   IOField "I/O field_72" at 566,349 size 60x22; Authorization "Parameter Change"; FormatPattern 9999
      ProcessValue <- "84_Setpoints_PIT402_Main_HighHigh"
   TextField "Text field_38" at 8,349 size 53x22; Text 'IW116'
   IOField "I/O field_29" at 566,511 size 60x22; FormatPattern 9999
   IOField "I/O field_30" at 499,511 size 60x22; FormatPattern 9999
   IOField "I/O field_32" at 361,552 size 60x22; FormatPattern 9999
   IOField "I/O field_33" at 429,552 size 60x22; FormatPattern 9999
   IOField "I/O field_34" at 565,552 size 60x22; FormatPattern 9999
   IOField "I/O field_35" at 498,552 size 60x22; FormatPattern 9999
   TextField "Text field_39" at 1109,687 size 151x62; Text 'To BC Analogue Inputs'
   AlarmView "Alarm view_1" at 0,777 size 1280x23
   TextField "Text field_40" at 23,309 size 1188x123; Text 'Re - Work Required Througout This page'
   Group "Group" at 455,41 size 373x50
   Button "HmiScreenItemData_8" at 469,45 size 355x40; TextOn 'Back'; TextOff 'Text'
   TextField "Screen title" at 455,41 size 373x50; Text 'Screen title'

screen "BC Analogue Outputs" 1280x800, template "Template"
   on GenerateScreen: "TitleUpdater"()
   Button "HmiScreenItemData_1" at 1,1 size 150x43; TextOn 'Back'; TextOff 'Commissioning'
      on Release: ActivateScreen("Commissioning Main Page", 0)
   Button "Button_15" at 34,732 size 100x35; TextOn 'BWTS Digital Inputs'; TextOff 'Back'
      on Click: ActivateScreen("BC Analogue Inputs", 0)
   AlarmView "Alarm view_1" at 0,777 size 1280x23
   TextField "Text field_90" at 750,328 size 64x20; Text 'Reading'
   TextField "Text field_41" at 553,328 size 89x20; Text 'Description'
   TextField "Text field_43" at 437,328 size 37x20; Text 'AO'
   TextField "Text field_52" at 437,295 size 364x26; Text 'Burner Control System PLC (Rack 2)'
   TextField "Text field_4" at 481,444 size 220x22; Text 'Main Fuel Reg Valve Control'
   IOField "I/O field_4" at 749,446 size 70x22; FormatPattern 9999; Unit %
      ProcessValue <- "16_AQ_Data_CV203_CNTRL"
   TextField "Text field_8" at 428,444 size 53x22; Text 'QW100'
   TextField "Text field_9" at 481,368 size 220x22; Text 'Spare'
   TextField "Text field_12" at 480,482 size 220x22; Text 'Main Atom Air Reg Valve Control'
   IOField "I/O field_5" at 749,481 size 70x22; FormatPattern 9999; Unit %
      ProcessValue <- "16_AQ_Data_CV111_CNTRL"
   TextField "Text field_13" at 427,482 size 53x22; Text 'QW102'
   Button "Button_7" at 716,442 size 29x26; TextOff '+'
      on Press: function_b14e0dd5("80_From_HMI_MAN_AQ_INC_100(1)", 0)
      Visibility <- "82_To_HMI_CRNT_MODE_IGG"
   Button "Button_8" at 824,442 size 29x26; TextOff '-'
      on Press: function_b14e0dd5("80_From_HMI_MAN_AQ_DEC_100(1)", 0)
      Visibility <- "82_To_HMI_CRNT_MODE_IGG"
   Button "Button_9" at 716,480 size 29x26; TextOff '+'
      on Press: function_b14e0dd5("80_From_HMI_MAN_AQ_INC_102", 0)
      Visibility <- "82_To_HMI_CRNT_MODE_IGG"
   Button "Button_10" at 824,480 size 29x26; TextOff '-'
      on Press: function_b14e0dd5("80_From_HMI_MAN_AQ_DEC_102", 0)
      Visibility <- "82_To_HMI_CRNT_MODE_IGG"
   Button "Button_11" at 716,364 size 29x26; TextOff '+'
      on Click: SetBit("80_From_HMI_MAN_AQ_INC_96")
      Visibility <- "82_To_HMI_CRNT_MODE_IGG"
   Button "Button_12" at 824,364 size 29x26; TextOff '-'
      on Click: SetBit("80_From_HMI_MAN_AQ_DEC_96")
      Visibility <- "82_To_HMI_CRNT_MODE_IGG"
   Button "Button_13" at 716,405 size 29x26; TextOff '+'
      on Click: SetBit("80_From_HMI_MAN_AQ_INC_98")
      Visibility <- "82_To_HMI_CRNT_MODE_IGG"
   Button "Button_14" at 824,405 size 29x26; TextOff '-'
      on Click: SetBit("80_From_HMI_MAN_AQ_DEC_98")
      Visibility <- "82_To_HMI_CRNT_MODE_IGG"
   IOField "I/O field_6" at 749,368 size 70x22; FormatPattern 9.9; Unit  
      ProcessValue <- "16_AQ_Data_R2_SPR_AQ_96"
   IOField "I/O field_7" at 749,408 size 70x22; FormatPattern 9.9; Unit  
      ProcessValue <- "16_AQ_Data_R2_SPR_AQ_98"
   TextField "Text field_14" at 481,408 size 220x22; Text 'Spare'
   TextField "Text field_15" at 429,368 size 53x22; Text 'QW96'
   TextField "Text field_16" at 428,408 size 53x22; Text 'QW98'
   Group "Group" at 455,41 size 373x50
   Button "HmiScreenItemData_8" at 469,45 size 355x40; TextOn 'Back'; TextOff 'Text'
   TextField "Screen title" at 455,41 size 373x50; Text 'Screen title'

screen "GCU Analogue Outputs" 1280x800, template "Template"
   on GenerateScreen: "TitleUpdater"()
   Button "HmiScreenItemData_1" at 1,1 size 150x43; TextOn 'Back'; TextOff 'Commissioning'
      on Release: ActivateScreen("Commissioning Main Page", 0)
   Button "Button_15" at 34,732 size 100x35; TextOn 'BWTS Digital Inputs'; TextOff 'Back'
      on Click: ActivateScreen("BC Analogue Inputs", 0)
   AlarmView "Alarm view_1" at 0,777 size 1280x23
   TextField "Text field_90" at 750,328 size 64x20; Text 'Reading'
   TextField "Text field_41" at 553,328 size 89x20; Text 'Description'
   TextField "Text field_43" at 437,328 size 37x20; Text 'AO'
   TextField "Text field_52" at 437,295 size 336x26; Text 'GCU Control System PLC (Rack 3)'
   TextField "Text field_4" at 481,444 size 220x22; Text 'Spare'
   IOField "I/O field_4" at 749,446 size 70x22; FormatPattern 9999
      ProcessValue <- "16_AQ_Data_R3_SPR_AQ_804"
   TextField "Text field_8" at 428,444 size 53x22; Text 'QW804'
   TextField "Text field_9" at 481,368 size 220x22; Text 'CV405 GAS VENT POSITION'
   TextField "Text field_12" at 480,482 size 220x22; Text 'Spare'
   IOField "I/O field_5" at 749,481 size 70x22; FormatPattern 9999
      ProcessValue <- "16_AQ_Data_R3_SPR_AQ_806"
   TextField "Text field_13" at 427,482 size 53x22; Text 'QW806'
   Button "Button_7" at 716,442 size 29x26; TextOff '+'
      on Press: function_b14e0dd5("80_From_HMI_MAN_AQ_INC_804", 0)
      Visibility <- "82_To_HMI_CRNT_MODE_GCU"
   Button "Button_8" at 824,442 size 29x26; TextOff '-'
      on Press: function_b14e0dd5("80_From_HMI_MAN_AQ_DEC_804", 0)
      Visibility <- "82_To_HMI_CRNT_MODE_GCU"
   Button "Button_9" at 717,480 size 29x26; TextOff '+'
      on Press: function_b14e0dd5("80_From_HMI_MAN_AQ_INC_806", 0)
      Visibility <- "82_To_HMI_CRNT_MODE_GCU"
   Button "Button_10" at 825,480 size 29x26; TextOff '-'
      on Press: function_b14e0dd5("80_From_HMI_MAN_AQ_DEC_806", 0)
      Visibility <- "82_To_HMI_CRNT_MODE_GCU"
   Button "Button_11" at 716,364 size 29x26; TextOff '+'
      Visibility <- "82_To_HMI_CRNT_MODE_GCU"
      on Press: function_b14e0dd5("80_From_HMI_MAN_AQ_INC_800", 0)
   Button "Button_12" at 824,364 size 29x26; TextOff '-'
      Visibility <- "82_To_HMI_CRNT_MODE_GCU"
      on Press: function_b14e0dd5("80_From_HMI_MAN_AQ_DEC_800", 0)
   Button "Button_13" at 717,405 size 29x26; TextOff '+'
      Visibility <- "82_To_HMI_CRNT_MODE_GCU"
      on Press: function_b14e0dd5("80_From_HMI_MAN_AQ_INC_802", 0)
   Button "Button_14" at 825,405 size 29x26; TextOff '-'
      Visibility <- "82_To_HMI_CRNT_MODE_GCU"
      on Press: function_b14e0dd5("80_From_HMI_MAN_AQ_DEC_802", 0)
   IOField "I/O field_6" at 750,368 size 70x22; FormatPattern 999; Unit   %
      ProcessValue <- "16_AQ_Data_CV405_CNTRL"
   IOField "I/O field_7" at 751,408 size 70x22; FormatPattern 9999; Unit  
      ProcessValue <- "16_AQ_Data_R3_SPR_AQ_802"
   TextField "Text field_14" at 481,408 size 220x22; Text 'Spare'
   TextField "Text field_15" at 429,368 size 53x22; Text 'QW800'
   TextField "Text field_16" at 428,408 size 53x22; Text 'QW802'
   Group "Group" at 455,41 size 373x50
   Button "HmiScreenItemData_8" at 469,45 size 355x40; TextOn 'Back'; TextOff 'Text'
   TextField "Screen title" at 455,41 size 373x50; Text 'Screen title'

screen "BWT Analogue Outputs" 1280x800, template "Template"
   on GenerateScreen: "TitleUpdater"()
   Button "HmiScreenItemData_1" at 1,1 size 150x43; TextOn 'Back'; TextOff 'Commissioning'
      on Release: ActivateScreen("Commissioning Main Page", 0)
   TextField "Text field_90" at 799,171 size 64x20; Text 'Reading'
   TextField "Text field_41" at 602,171 size 89x20; Text 'Description'
   TextField "Text field_43" at 486,171 size 37x20; Text 'AO'
   TextField "Text field_52" at 486,138 size 340x26; Text 'BWT Control System PLC (Rack 3)'
   TextField "Text field_4" at 530,287 size 220x22; Text 'Main Fuel Reg Valve Control'
   IOField "I/O field_4" at 798,289 size 70x22; FormatPattern 9999; Unit %
      ProcessValue <- "16_AQ_Data_CV203_CNTRL"
   TextField "Text field_8" at 477,287 size 53x22; Text 'QW100'
   TextField "Text field_9" at 530,211 size 220x22; Text 'Spare'
   TextField "Text field_12" at 529,325 size 220x22; Text 'Main Atom Air Reg Valve Control'
   IOField "I/O field_5" at 798,324 size 70x22; FormatPattern 9999; Unit %
      ProcessValue <- "16_AQ_Data_CV111_CNTRL"
   TextField "Text field_13" at 476,325 size 53x22; Text 'QW102'
   Button "Button_7" at 765,285 size 29x26; TextOff '+'
      on Press: function_b14e0dd5("80_From_HMI_MAN_AQ_INC_100(1)", 0)
      Visibility <- "82_To_HMI_CRNT_MODE_IGG"
   Button "Button_8" at 873,285 size 29x26; TextOff '-'
      on Press: function_b14e0dd5("80_From_HMI_MAN_AQ_DEC_100(1)", 0)
      Visibility <- "82_To_HMI_CRNT_MODE_IGG"
   Button "Button_9" at 766,323 size 29x26; TextOff '+'
      on Press: function_b14e0dd5("80_From_HMI_MAN_AQ_INC_102", 0)
      Visibility <- "82_To_HMI_CRNT_MODE_IGG"
   Button "Button_10" at 874,323 size 29x26; TextOff '-'
      on Press: function_b14e0dd5("80_From_HMI_MAN_AQ_DEC_102", 0)
      Visibility <- "82_To_HMI_CRNT_MODE_IGG"
   Button "Button_11" at 765,207 size 29x26; TextOff '+'
      on Click: SetBit("80_From_HMI_MAN_AQ_INC_96")
      Visibility <- "82_To_HMI_CRNT_MODE_IGG"
   Button "Button_12" at 873,207 size 29x26; TextOff '-'
      on Click: SetBit("80_From_HMI_MAN_AQ_DEC_96")
      Visibility <- "82_To_HMI_CRNT_MODE_IGG"
   Button "Button_13" at 766,248 size 29x26; TextOff '+'
      on Click: SetBit("80_From_HMI_MAN_AQ_INC_98")
      Visibility <- "82_To_HMI_CRNT_MODE_IGG"
   Button "Button_14" at 874,248 size 29x26; TextOff '-'
      on Click: SetBit("80_From_HMI_MAN_AQ_DEC_98")
      Visibility <- "82_To_HMI_CRNT_MODE_IGG"
   IOField "I/O field_6" at 799,211 size 70x22; FormatPattern 9.9; Unit  
      ProcessValue <- "16_AQ_Data_R2_SPR_AQ_96"
   IOField "I/O field_7" at 800,251 size 70x22; FormatPattern 9.9; Unit  
      ProcessValue <- "16_AQ_Data_R2_SPR_AQ_98"
   TextField "Text field_14" at 530,251 size 220x22; Text 'Spare'
   TextField "Text field_15" at 478,211 size 53x22; Text 'QW96'
   TextField "Text field_16" at 477,251 size 53x22; Text 'QW98'
   Button "Button_15" at 34,732 size 100x35; TextOn 'BWTS Digital Inputs'; TextOff 'Back'
      on Click: ActivateScreen("BC Analogue Inputs", 0)
   AlarmView "Alarm view_1" at 0,777 size 1280x23
   TextField "Text field_1" at 23,309 size 1188x123; Text 'Re - Work Required Througout This page'
   Group "Group" at 455,41 size 373x50
   Button "HmiScreenItemData_8" at 469,45 size 355x40; TextOn 'Back'; TextOff 'Text'
   TextField "Screen title" at 455,41 size 373x50; Text 'Screen title'

screen "BC Target Setpoints" 1280x800, template "Template"
   on GenerateScreen: "TitleUpdater"()
   Button "HmiScreenItemData_1" at 1,1 size 150x43; TextOn 'Back'; TextOff 'Commissioning'
      on Release: ActivateScreen("Commissioning Main Page", 0)
   AlarmView "Alarm view_1" at 0,777 size 1280x23
   TextField "Text field_25" at 394,430 size 407x22; Text 'PIT-113: IGG Main Atom Air Pressure Target'
   TextField "Text field_29" at 814,210 size 68x20; Text 'Setpoint'
   TextField "Text field_33" at 393,468 size 408x22; Text 'PIT-205: IGG Main Fuel Pressure Target'
   IOField "I/O field_58" at 816,468 size 60x22; Authorization "Parameter Change"; FormatPattern 999.99
      ProcessValue <- "84_Setpoints_PIT205_Target(1)"
   TextField "Text field_35" at 394,552 size 406x22; Text 'E-600: O2 Cargo Blanketing Target'
   TextField "Text field_65" at 394,236 size 411x22; Text 'PIT-402: IG Outlet Pressure Pilot Target'
   TextField "Text field_67" at 394,274 size 410x22; Text 'PIT-402: IG Outlet Pressure Main Target'
   TextField "Text field_69" at 395,313 size 407x22; Text 'PIT-402: IG Outlet Pressure Post Target Start'
   TextField "Text field_71" at 395,352 size 406x22; Text 'PIT-402: IG Outlet Pressure Post Target Maximum'
   TextField "Text field_73" at 395,391 size 407x22; Text 'FD-001: Igniter Target'
   TextField "Text field_42" at 394,210 size 89x20; Text 'Description'
   IOField "I/O field_128" at 816,236 size 60x22; Authorization "Parameter Change"; FormatPattern 999.9
      ProcessValue <- "84_Setpoints_PIT402_Pilot_Target(1)"
   IOField "I/O field_133" at 816,274 size 60x22; Authorization "Parameter Change"; FormatPattern 999.9
      ProcessValue <- "84_Setpoints_PIT402_Main_Target(1)"
   IOField "I/O field_138" at 816,313 size 60x22; Authorization "Parameter Change"; FormatPattern 999.9
      ProcessValue <- "84_Setpoints_PIT402_Post_Target_Start"
   IOField "I/O field_53" at 816,430 size 60x22; Authorization "Parameter Change"; FormatPattern 999.9
      ProcessValue <- "84_Setpoints_PIT113_Pilot_Target(1)"
   IOField "I/O field_148" at 816,391 size 60x22; Authorization "Parameter Change"; FormatPattern 999.9
      ProcessValue <- "84_Setpoints_FD001_Min"
   IOField "I/O field_64" at 816,552 size 60x22; Authorization "Parameter Change"; FormatPattern 99.9
      ProcessValue <- "84_Setpoints_E600_CB_Target"
   TextField "Text field_53" at 393,184 size 213x26; Text 'IGG Target Setpoints'
   IOField "I/O field_5" at 815,352 size 60x22; Authorization "Parameter Change"; FormatPattern 999.9
      ProcessValue <- "84_Setpoints_PIT401_Post_Target_Max"
   TextField "Text field_1" at 394,510 size 406x22; Text 'E-600: O2 Ballast Water Treatment Target'
   IOField "I/O field_2" at 816,510 size 60x22; Authorization "Parameter Change"; FormatPattern 9.99
      ProcessValue <- "84_Setpoints_E600_BWT_Target"
   TextField "Text field_2" at 394,595 size 406x22; Text 'PIT-402 Target Ramp Time (s)'
   IOField "I/O field_1" at 816,595 size 60x22; Authorization "Parameter Change"; FormatPattern 99
      ProcessValue <- "19_AUTO_CMNDS_Data_PIT402_Target"
   Group "Group" at 455,41 size 373x50
   Button "HmiScreenItemData_8" at 469,45 size 355x40; TextOn 'Back'; TextOff 'Text'
   TextField "Screen title" at 455,41 size 373x50; Text 'Screen title'

screen "BC Process Times" 1280x800, template "Template"
   on GenerateScreen: "TitleUpdater"()
   Button "HmiScreenItemData_1" at 1,1 size 150x43; TextOn 'Back'; TextOff 'Commissioning'
      on Release: ActivateScreen("Commissioning Main Page", 0)
   Button "Button_1" at 21,736 size 161x32; TextOff 'IGG Step Times'
      on Activate: ActivateScreen("IGG Max Step Times", 0)
   Button "Button_2" at 1091,736 size 161x32; TextOff 'BC Step Times'
      on Activate: ActivateScreen("BC Max Step Times", 0)
   AlarmView "Alarm view_1" at 0,777 size 1280x23
   TextField "Text field_2" at 262,326 size 271x22; Text 'CV114 Open Delay Time'
   TextField "Text field_3" at 551,161 size 65x20; Text 'Time (s)'
   TextField "Text field_4" at 262,354 size 273x22; Text 'CV206 Open Delay Time'
   IOField "I/O field_1" at 546,354 size 60x22; Authorization "Parameter Change"; FormatPattern 999
      ProcessValue <- "86_Times_CV206_OPEN_TIME"
   TextField "Text field_5" at 262,411 size 270x22; Text 'CV215 Open Delay Time'
   TextField "Text field_6" at 262,186 size 272x22; Text 'CV127 Open #1 Delay Time'
   TextField "Text field_7" at 262,214 size 272x22; Text 'CV127 Closed Delay Time'
   TextField "Text field_8" at 262,242 size 271x22; Text 'CV127 Open #2 Delay Time'
   TextField "Text field_9" at 262,270 size 270x22; Text 'CV124 Open Delay Time'
   TextField "Text field_10" at 262,298 size 270x22; Text 'CV124 Close Delay Purge Time'
   TextField "Text field_11" at 262,161 size 89x20; Text 'Description'
   IOField "I/O field_3" at 546,186 size 60x22; Authorization "Parameter Change"; FormatPattern 999
      ProcessValue <- "86_Times_CV127_OPEN_TIME_#1"
   IOField "I/O field_4" at 546,214 size 60x22; Authorization "Parameter Change"; FormatPattern 999
      ProcessValue <- "86_Times_CV127_CLOSED_TIME"
   IOField "I/O field_6" at 546,242 size 60x22; Authorization "Parameter Change"; FormatPattern 999
      ProcessValue <- "86_Times_CV127_OPEN_TIME_#2"
   IOField "I/O field_8" at 546,298 size 60x22; Authorization "Parameter Change"; FormatPattern 999
      ProcessValue <- "86_Times_CV124_CLOSE_TIME_PRG"
   IOField "I/O field_9" at 546,410 size 60x22; Authorization "Parameter Change"; FormatPattern 999
      ProcessValue <- "86_Times_CV215_OPEN_TIME"
   TextField "Text field_12" at 261,135 size 178x26; Text 'BC Process Times'
   IOField "I/O field_10" at 546,270 size 60x22; Authorization "Parameter Change"; FormatPattern 999
      ProcessValue <- "86_Times_CV124_OPEN_TIME"
   TextField "Text field_13" at 262,383 size 270x22; Text 'CV207 Open Delay Time'
   IOField "I/O field_11" at 546,382 size 60x22; Authorization "Parameter Change"; FormatPattern 999
      ProcessValue <- "86_Times_CV207_OPEN_TIME"
   TextField "Text field_17" at 262,439 size 270x22; Text 'CV215 Close Delay Purge Time'
   IOField "I/O field_16" at 546,438 size 60x22; Authorization "Parameter Change"; FormatPattern 999
      ProcessValue <- "86_Times_CV215_CLOSE_TIME_PRG"
   TextField "Text field_18" at 262,467 size 270x22; Text 'CV216 Open Delay Time'
   IOField "I/O field_17" at 546,466 size 60x22; Authorization "Parameter Change"; FormatPattern 999
      ProcessValue <- "86_Times_CV216_OPEN_TIME"
   TextField "Text field_19" at 262,495 size 269x22; Text 'CV216 Close Delay Purge Time'
   IOField "I/O field_18" at 546,494 size 60x22; Authorization "Parameter Change"; FormatPattern 999
      ProcessValue <- "86_Times_CV216_CLOSE_TIME_PRG"
   TextField "Text field_20" at 262,523 size 269x22; Text 'CV216 Open Delay Purge Time'
   IOField "I/O field_19" at 546,522 size 60x22; Authorization "Parameter Change"; FormatPattern 999
      ProcessValue <- "86_Times_CV216_OPEN_TIME_PRG"
   TextField "Text field_21" at 262,552 size 269x22; Text 'CV206 Close Delay Time'
   IOField "I/O field_20" at 546,551 size 60x22; Authorization "Parameter Change"; FormatPattern 999
      ProcessValue <- "86_Times_CV206_CLOSE_TIME"
   TextField "Text field_22" at 636,186 size 269x22; Text 'CV207 Close Delay Time'
   IOField "I/O field_21" at 916,186 size 60x22; Authorization "Parameter Change"; FormatPattern 999
      ProcessValue <- "86_Times_CV207_CLOSE_TIME"
   TextField "Text field_23" at 636,160 size 89x20; Text 'Description'
   TextField "Text field_24" at 923,161 size 65x20; Text 'Time (s)'
   TextField "Text field_26" at 636,214 size 269x22; Text 'CV114 Close Delay Time'
   IOField "I/O field_22" at 916,214 size 60x22; Authorization "Parameter Change"; FormatPattern 999
      ProcessValue <- "86_Times_CV114_CLOSE_TIME"
   TextField "Text field_27" at 636,242 size 269x22; Text 'CV215 Close Delay Time'
   IOField "I/O field_23" at 916,242 size 60x22; Authorization "Parameter Change"; FormatPattern 999
      ProcessValue <- "86_Times_CV215_CLOSE_TIME"
   TextField "Text field_28" at 636,270 size 269x22; Text 'CV216 Close Delay Time'
   IOField "I/O field_24" at 916,270 size 60x22; Authorization "Parameter Change"; FormatPattern 999
      ProcessValue <- "86_Times_CV216_CLOSE_TIME"
   TextField "Text field_30" at 636,298 size 269x22; Text 'CV124 Close Delay Time'
   IOField "I/O field_25" at 916,298 size 60x22; Authorization "Parameter Change"; FormatPattern 999
      ProcessValue <- "86_Times_CV124_CLOSE_TIME"
   TextField "Text field_31" at 636,326 size 269x22; Text 'X001 Maximum Run Time'
   IOField "I/O field_26" at 916,326 size 60x22; Authorization "Parameter Change"; FormatPattern 999
      ProcessValue <- "86_Times_X001_MAX_RUN_TIME"
   TextField "Text field_32" at 636,354 size 269x22; Text 'X001 Run Confirmation Time'
   IOField "I/O field_27" at 916,354 size 60x22; Authorization "Parameter Change"; FormatPattern 999
      ProcessValue <- "86_Times_X001_RUN_CNF_TIME"
   TextField "Text field_34" at 636,383 size 269x22; Text 'Flame Detection Delay'
   IOField "I/O field_28" at 916,382 size 60x22; Authorization "Parameter Change"; FormatPattern 999
      ProcessValue <- "86_Times_FD_DET_DELAY"
   TextField "Text field_36" at 636,411 size 269x22; Text 'Flame Verification Time'
   IOField "I/O field_29" at 916,410 size 60x22; Authorization "Parameter Change"; FormatPattern 999
      ProcessValue <- "86_Times_FD_VRFCTN_TIME"
   TextField "Text field_37" at 636,439 size 269x22; Text 'Flame Detection Time'
   IOField "I/O field_30" at 916,438 size 60x22; Authorization "Parameter Change"; FormatPattern 999
      ProcessValue <- "86_Times_FDU_DET_TIME"
   TextField "Text field_38" at 636,467 size 269x22; Text 'Max Ignition Sequence Run Time'
   IOField "I/O field_31" at 916,466 size 60x22; Authorization "Parameter Change"; FormatPattern 999
      ProcessValue <- "86_Times_MAX_IGNTN_SEQ_TIME"
   TextField "Text field_39" at 636,495 size 269x22; Text 'Max Main Burner Sequence Run Time'
      Visibility <- "AlwaysTRUE"
   IOField "I/O field_32" at 916,494 size 60x22; Authorization "Parameter Change"; FormatPattern 999; Unit h
      ProcessValue <- "86_Times_MAX_MAIN_BURN_SEQ_TIME"
      Visibility <- "AlwaysTRUE"
   TextField "Text field_40" at 636,523 size 269x22; Text 'Max Pilot Burner Purge Sequence Run Time'
   IOField "I/O field_33" at 916,522 size 60x22; Authorization "Parameter Change"; FormatPattern 999
      ProcessValue <- "86_Times_MAX_PILOT_PURGE_SEQ_TIME"
   TextField "Text field_41" at 636,552 size 269x22; Text 'O2 Check Delay Time'
   IOField "I/O field_34" at 916,551 size 60x22; Authorization "Parameter Change"; FormatPattern 999
      ProcessValue <- "86_Times_O2_CHECK_TIME"
   IOField "I/O field_7" at 546,326 size 60x22; Authorization "Parameter Change"; FormatPattern 999
      ProcessValue <- "86_Times_CV114_OPEN_TIME"
   TextField "Text field_43" at 636,582 size 269x22; Text 'Flame Fail Delay'
   IOField "I/O field_35" at 916,581 size 60x22; Authorization "Parameter Change"; FormatPattern 999
      ProcessValue <- "80_From_HMI_FLM_FAIL_DLY"
   Switch "Switch_1" at 987,492 size 32x29; CaptionText 'Switch'; TextOn 'ON'; TextOff 'OFF'; Authorization "User administration"; PictureOff "Design_5_PilotLight_Green_Off"; PictureOn "Design_5_PilotLight_Green_On"
      on Activate: SetBit("80_From_HMI_BurnerProgramedStop")
      ProcessValue <- "80_From_HMI_BurnerProgramedStop"
      Visibility <- "AlwaysTRUE"
   TextField "Text field_44" at 636,613 size 269x22; Text 'FS317 Delayed Fault'
   IOField "I/O field_36" at 916,613 size 60x22; Authorization "Parameter Change"; FormatPattern 999
      ProcessValue <- "86_Times_FS317 delay"
   TextField "Text field_45" at 636,644 size 269x22; Text 'FS320 Delayed Fault'
   IOField "I/O field_37" at 916,644 size 60x22; Authorization "Parameter Change"; FormatPattern 999
      ProcessValue <- "86_Times_FS320 delay"
   TextField "Text field_46" at 262,581 size 269x22; Text 'FS359 Delayed Fault'
   IOField "I/O field_38" at 546,581 size 60x22; Authorization "Parameter Change"; FormatPattern 999
      ProcessValue <- "80_From_HMI_PIT 359 delay"
   TextField "Text field_47" at 262,612 size 269x22; Text 'FS316 Delayed Fault'
   IOField "I/O field_39" at 546,612 size 60x22; Authorization "Parameter Change"; FormatPattern 999
      ProcessValue <- "80_From_HMI_PIT 316 delay"
   Group "Group" at 455,41 size 373x50
   TextField "Text field_1" at 262,643 size 269x22; Text 'PS101 Delayed Fault'
   IOField "I/O field_2" at 546,643 size 60x22; Authorization "Parameter Change"; FormatPattern 999
      ProcessValue <- "86_Times_PS101 Alarm Delay"
   Button "HmiScreenItemData_8" at 469,45 size 355x40; TextOn 'Back'; TextOff 'Text'
   TextField "Screen title" at 455,41 size 373x50; Text 'Screen title'

screen "GCU Max Step Times" 1280x800, template "Template"
   on GenerateScreen: "TitleUpdater"()
   Button "HmiScreenItemData_1" at 1,1 size 150x43; TextOn 'Back'; TextOff 'Commissioning'
      on Release: ActivateScreen("Commissioning Main Page", 0)
   TextField "Text field_29" at 130,95 size 75x25; Text 'Time (ms)'
   TextField "Text field_65" at 40,130 size 75x25; Text 'Step 001'
   TextField "Text field_42" at 40,95 size 75x25; Text 'STEP'
   IOField "I/O field_128" at 130,130 size 75x25; Authorization "Parameter Change"; FormatPattern 999999
      ProcessValue <- "86_Times_STEP_MAX_TIME_STP_001"
   TextField "Text field_53" at 40,66 size 262x26; Text 'GCU Maximum Step Times'
   TextField "Text field_1" at 385,95 size 75x25; Text 'Time (ms)'
   TextField "Text field_2" at 295,130 size 75x25; Text 'Step 170'
   TextField "Text field_3" at 295,95 size 75x25; Text 'STEP'
   IOField "I/O field_1" at 385,130 size 75x25; Authorization "Parameter Change"; FormatPattern 999999
      ProcessValue <- "86_Times_STEP_MAX_TIME_STP_170"
   TextField "Text field_4" at 640,95 size 75x25; Text 'Time (ms)'
   TextField "Text field_5" at 550,130 size 75x25; Text 'Step 350'
   TextField "Text field_6" at 550,95 size 75x25; Text 'STEP'
   IOField "I/O field_2" at 640,130 size 75x25; Authorization "Parameter Change"; FormatPattern 999999
      ProcessValue <- "86_Times_STEP_MAX_TIME_STP_350"
   TextField "Text field_7" at 895,95 size 75x25; Text 'Time (ms)'
   TextField "Text field_8" at 805,130 size 75x25; Text 'Step 530'
   TextField "Text field_9" at 805,95 size 75x25; Text 'STEP'
   IOField "I/O field_3" at 895,130 size 75x25; Authorization "Parameter Change"; FormatPattern 999999
      ProcessValue <- "86_Times_STEP_MAX_TIME_STP_530"
   TextField "Text field_10" at 1150,95 size 75x25; Text 'Time (ms)'
   TextField "Text field_12" at 1060,95 size 75x25; Text 'STEP'
   TextField "Text field_13" at 40,165 size 75x25; Text 'Step 005'
   IOField "I/O field_5" at 130,165 size 75x25; Authorization "Parameter Change"; FormatPattern 999999
      ProcessValue <- "86_Times_STEP_MAX_TIME_STP_005"
   TextField "Text field_14" at 295,165 size 75x25; Text 'Step 180'
   IOField "I/O field_6" at 385,165 size 75x25; Authorization "Parameter Change"; FormatPattern 999999
      ProcessValue <- "86_Times_STEP_MAX_TIME_STP_180"
   TextField "Text field_15" at 550,165 size 75x25; Text 'Step 360'
   IOField "I/O field_7" at 640,165 size 75x25; Authorization "Parameter Change"; FormatPattern 999999
      ProcessValue <- "86_Times_STEP_MAX_TIME_STP_360"
   TextField "Text field_16" at 805,165 size 75x25; Text 'Step 540'
   IOField "I/O field_8" at 895,165 size 75x25; Authorization "Parameter Change"; FormatPattern 999999
      ProcessValue <- "86_Times_STEP_MAX_TIME_STP_540"
   TextField "Text field_18" at 40,200 size 75x25; Text 'Step 010'
   IOField "I/O field_10" at 130,200 size 75x25; Authorization "Parameter Change"; FormatPattern 999999
      ProcessValue <- "86_Times_STEP_MAX_TIME_STP_010"
   TextField "Text field_19" at 295,200 size 75x25; Text 'Step 190'
   IOField "I/O field_11" at 385,200 size 75x25; Authorization "Parameter Change"; FormatPattern 999999
      ProcessValue <- "86_Times_STEP_MAX_TIME_STP_190"
   TextField "Text field_20" at 550,200 size 75x25; Text 'Step 370'
   IOField "I/O field_12" at 640,200 size 75x25; Authorization "Parameter Change"; FormatPattern 999999
      ProcessValue <- "86_Times_STEP_MAX_TIME_STP_370"
   TextField "Text field_21" at 805,200 size 75x25; Text 'Step 550'
   IOField "I/O field_13" at 895,200 size 75x25; Authorization "Parameter Change"; FormatPattern 999999
      ProcessValue <- "86_Times_STEP_MAX_TIME_STP_550"
   TextField "Text field_23" at 40,235 size 75x25; Text 'Step 020'
   IOField "I/O field_15" at 130,235 size 75x25; Authorization "Parameter Change"; FormatPattern 999999
      ProcessValue <- "86_Times_STEP_MAX_TIME_STP_020"
   TextField "Text field_24" at 295,235 size 75x25; Text 'Step 200'
   IOField "I/O field_16" at 385,235 size 75x25; Authorization "Parameter Change"; FormatPattern 999999
      ProcessValue <- "86_Times_STEP_MAX_TIME_STP_200"
   TextField "Text field_25" at 550,235 size 75x25; Text 'Step 380'
   IOField "I/O field_17" at 640,235 size 75x25; Authorization "Parameter Change"; FormatPattern 999999
      ProcessValue <- "86_Times_STEP_MAX_TIME_STP_380"
   TextField "Text field_26" at 805,235 size 75x25; Text 'Step 560'
   IOField "I/O field_18" at 895,235 size 75x25; Authorization "Parameter Change"; FormatPattern 999999
      ProcessValue <- "86_Times_STEP_MAX_TIME_STP_560"
   TextField "Text field_28" at 40,270 size 75x25; Text 'Step 030'
   IOField "I/O field_20" at 130,270 size 75x25; Authorization "Parameter Change"; FormatPattern 999999
      ProcessValue <- "86_Times_STEP_MAX_TIME_STP_030"
   TextField "Text field_30" at 295,270 size 75x25; Text 'Step 210'
   IOField "I/O field_21" at 385,270 size 75x25; Authorization "Parameter Change"; FormatPattern 999999
      ProcessValue <- "86_Times_STEP_MAX_TIME_STP_210"
   TextField "Text field_31" at 550,270 size 75x25; Text 'Step 390'
   IOField "I/O field_22" at 640,270 size 75x25; Authorization "Parameter Change"; FormatPattern 999999
      ProcessValue <- "86_Times_STEP_MAX_TIME_STP_390"
   TextField "Text field_32" at 805,270 size 75x25; Text 'Step 570'
   IOField "I/O field_23" at 895,270 size 75x25; Authorization "Parameter Change"; FormatPattern 999999
      ProcessValue <- "86_Times_STEP_MAX_TIME_STP_570"
   TextField "Text field_34" at 40,305 size 75x25; Text 'Step 040'
   IOField "I/O field_25" at 130,305 size 75x25; Authorization "Parameter Change"; FormatPattern 999999
      ProcessValue <- "86_Times_STEP_MAX_TIME_STP_040"
   TextField "Text field_35" at 295,305 size 75x25; Text 'Step 220'
   IOField "I/O field_26" at 385,305 size 75x25; Authorization "Parameter Change"; FormatPattern 999999
      ProcessValue <- "86_Times_STEP_MAX_TIME_STP_220"
   TextField "Text field_36" at 550,305 size 75x25; Text 'Step 400'
   IOField "I/O field_27" at 640,305 size 75x25; Authorization "Parameter Change"; FormatPattern 999999
      ProcessValue <- "86_Times_STEP_MAX_TIME_STP_400"
   TextField "Text field_37" at 805,305 size 75x25; Text 'Step 580'
   IOField "I/O field_28" at 895,305 size 75x25; Authorization "Parameter Change"; FormatPattern 999999
      ProcessValue <- "86_Times_STEP_MAX_TIME_STP_580"
   TextField "Text field_39" at 40,340 size 75x25; Text 'Step 050'
   IOField "I/O field_30" at 130,340 size 75x25; Authorization "Parameter Change"; FormatPattern 999999
      ProcessValue <- "86_Times_STEP_MAX_TIME_STP_050"
   TextField "Text field_40" at 295,340 size 75x25; Text 'Step 230'
   IOField "I/O field_31" at 385,340 size 75x25; Authorization "Parameter Change"; FormatPattern 999999
      ProcessValue <- "86_Times_STEP_MAX_TIME_STP_230"
   TextField "Text field_41" at 550,340 size 75x25; Text 'Step 410'
   IOField "I/O field_32" at 640,340 size 75x25; Authorization "Parameter Change"; FormatPattern 999999
      ProcessValue <- "86_Times_STEP_MAX_TIME_STP_410"
   TextField "Text field_43" at 805,340 size 75x25; Text 'Step 590'
   IOField "I/O field_33" at 895,340 size 75x25; Authorization "Parameter Change"; FormatPattern 999999
      ProcessValue <- "86_Times_STEP_MAX_TIME_STP_590"
   TextField "Text field_45" at 40,375 size 75x25; Text 'Step 060'
   IOField "I/O field_35" at 130,375 size 75x25; Authorization "Parameter Change"; FormatPattern 999999
      ProcessValue <- "86_Times_STEP_MAX_TIME_STP_060"
   TextField "Text field_46" at 295,375 size 75x25; Text 'Step 240'
   IOField "I/O field_36" at 385,375 size 75x25; Authorization "Parameter Change"; FormatPattern 999999
      ProcessValue <- "86_Times_STEP_MAX_TIME_STP_240"
   TextField "Text field_47" at 550,375 size 75x25; Text 'Step 420'
   IOField "I/O field_37" at 640,375 size 75x25; Authorization "Parameter Change"; FormatPattern 999999
      ProcessValue <- "86_Times_STEP_MAX_TIME_STP_420"
   TextField "Text field_48" at 805,375 size 75x25; Text 'Step 600'
   IOField "I/O field_38" at 895,375 size 75x25; Authorization "Parameter Change"; FormatPattern 999999
      ProcessValue <- "86_Times_STEP_MAX_TIME_STP_600"
   TextField "Text field_50" at 40,410 size 75x25; Text 'Step 070'
   IOField "I/O field_40" at 130,410 size 75x25; Authorization "Parameter Change"; FormatPattern 999999
      ProcessValue <- "86_Times_STEP_MAX_TIME_STP_070"
   TextField "Text field_51" at 295,410 size 75x25; Text 'Step 250'
   IOField "I/O field_41" at 385,410 size 75x25; Authorization "Parameter Change"; FormatPattern 999999
      ProcessValue <- "86_Times_STEP_MAX_TIME_STP_250"
   TextField "Text field_52" at 550,410 size 75x25; Text 'Step 430'
   IOField "I/O field_42" at 640,410 size 75x25; Authorization "Parameter Change"; FormatPattern 999999
      ProcessValue <- "86_Times_STEP_MAX_TIME_STP_430"
   TextField "Text field_54" at 805,410 size 75x25; Text 'Step 610'
   IOField "I/O field_43" at 895,410 size 75x25; Authorization "Parameter Change"; FormatPattern 999999
      ProcessValue <- "86_Times_STEP_MAX_TIME_STP_610"
   TextField "Text field_56" at 40,445 size 75x25; Text 'Step 080'
   IOField "I/O field_45" at 130,445 size 75x25; Authorization "Parameter Change"; FormatPattern 999999
      ProcessValue <- "86_Times_STEP_MAX_TIME_STP_080"
   TextField "Text field_57" at 295,445 size 75x25; Text 'Step 260'
   IOField "I/O field_46" at 385,445 size 75x25; Authorization "Parameter Change"; FormatPattern 999999
      ProcessValue <- "86_Times_STEP_MAX_TIME_STP_260"
   TextField "Text field_58" at 550,445 size 75x25; Text 'Step 440'
   IOField "I/O field_47" at 640,445 size 75x25; Authorization "Parameter Change"; FormatPattern 999999
      ProcessValue <- "86_Times_STEP_MAX_TIME_STP_440"
   TextField "Text field_59" at 805,445 size 75x25; Text 'Step 620'
   IOField "I/O field_48" at 895,445 size 75x25; Authorization "Parameter Change"; FormatPattern 999999
      ProcessValue <- "86_Times_STEP_MAX_TIME_STP_620"
   TextField "Text field_61" at 40,480 size 75x25; Text 'Step 090'
   IOField "I/O field_50" at 130,480 size 75x25; Authorization "Parameter Change"; FormatPattern 999999
      ProcessValue <- "86_Times_STEP_MAX_TIME_STP_090"
   TextField "Text field_62" at 295,480 size 75x25; Text 'Step 270'
   IOField "I/O field_51" at 385,480 size 75x25; Authorization "Parameter Change"; FormatPattern 999999
      ProcessValue <- "86_Times_STEP_MAX_TIME_STP_270"
   TextField "Text field_63" at 550,480 size 75x25; Text 'Step 450'
   IOField "I/O field_52" at 640,480 size 75x25; Authorization "Parameter Change"; FormatPattern 999999
      ProcessValue <- "86_Times_STEP_MAX_TIME_STP_450"
   TextField "Text field_64" at 805,480 size 75x25; Text 'Step 630'
   IOField "I/O field_53" at 895,480 size 75x25; Authorization "Parameter Change"; FormatPattern 999999
      ProcessValue <- "86_Times_STEP_MAX_TIME_STP_630"
   TextField "Text field_67" at 40,515 size 75x25; Text 'Step 100'
   IOField "I/O field_55" at 130,515 size 75x25; Authorization "Parameter Change"; FormatPattern 999999
      ProcessValue <- "86_Times_STEP_MAX_TIME_STP_100"
   TextField "Text field_68" at 295,515 size 75x25; Text 'Step 280'
   IOField "I/O field_56" at 385,515 size 75x25; Authorization "Parameter Change"; FormatPattern 999999
      ProcessValue <- "86_Times_STEP_MAX_TIME_STP_280"
   TextField "Text field_69" at 550,515 size 75x25; Text 'Step 460'
   IOField "I/O field_57" at 640,515 size 75x25; Authorization "Parameter Change"; FormatPattern 999999
      ProcessValue <- "86_Times_STEP_MAX_TIME_STP_460"
   TextField "Text field_72" at 40,550 size 75x25; Text 'Step 110'
   IOField "I/O field_60" at 130,550 size 75x25; Authorization "Parameter Change"; FormatPattern 999999
      ProcessValue <- "86_Times_STEP_MAX_TIME_STP_110"
   TextField "Text field_73" at 295,550 size 75x25; Text 'Step 290'
   IOField "I/O field_61" at 385,550 size 75x25; Authorization "Parameter Change"; FormatPattern 999999
      ProcessValue <- "86_Times_STEP_MAX_TIME_STP_290"
   TextField "Text field_74" at 550,550 size 75x25; Text 'Step 470'
   IOField "I/O field_62" at 640,550 size 75x25; Authorization "Parameter Change"; FormatPattern 999999
      ProcessValue <- "86_Times_STEP_MAX_TIME_STP_470"
   TextField "Text field_77" at 40,585 size 75x25; Text 'Step 120'
   IOField "I/O field_65" at 130,585 size 75x25; Authorization "Parameter Change"; FormatPattern 999999
      ProcessValue <- "86_Times_STEP_MAX_TIME_STP_120"
   TextField "Text field_78" at 295,585 size 75x25; Text 'Step 300'
   IOField "I/O field_66" at 385,585 size 75x25; Authorization "Parameter Change"; FormatPattern 999999
      ProcessValue <- "86_Times_STEP_MAX_TIME_STP_300"
   TextField "Text field_79" at 550,585 size 75x25; Text 'Step 480'
   IOField "I/O field_67" at 640,585 size 75x25; Authorization "Parameter Change"; FormatPattern 999999
      ProcessValue <- "86_Times_STEP_MAX_TIME_STP_480"
   TextField "Text field_82" at 40,620 size 75x25; Text 'Step 130'
   IOField "I/O field_70" at 130,620 size 75x25; Authorization "Parameter Change"; FormatPattern 999999
      ProcessValue <- "86_Times_STEP_MAX_TIME_STP_130"
   TextField "Text field_83" at 295,620 size 75x25; Text 'Step 310'
   IOField "I/O field_71" at 385,620 size 75x25; Authorization "Parameter Change"; FormatPattern 999999
      ProcessValue <- "86_Times_STEP_MAX_TIME_STP_310"
   TextField "Text field_84" at 550,620 size 75x25; Text 'Step 490'
   IOField "I/O field_72" at 640,620 size 75x25; Authorization "Parameter Change"; FormatPattern 999999
      ProcessValue <- "86_Times_STEP_MAX_TIME_STP_490"
   TextField "Text field_87" at 40,655 size 75x25; Text 'Step 140'
   IOField "I/O field_75" at 130,655 size 75x25; Authorization "Parameter Change"; FormatPattern 999999
      ProcessValue <- "86_Times_STEP_MAX_TIME_STP_140"
   TextField "Text field_88" at 295,655 size 75x25; Text 'Step 320'
   IOField "I/O field_76" at 385,655 size 75x25; Authorization "Parameter Change"; FormatPattern 999999
      ProcessValue <- "86_Times_STEP_MAX_TIME_STP_320"
   TextField "Text field_89" at 550,655 size 75x25; Text 'Step 500'
   IOField "I/O field_77" at 640,655 size 75x25; Authorization "Parameter Change"; FormatPattern 999999
      ProcessValue <- "86_Times_STEP_MAX_TIME_STP_500"
   TextField "Text field_92" at 40,690 size 75x25; Text 'Step 150'
   IOField "I/O field_80" at 130,690 size 75x25; Authorization "Parameter Change"; FormatPattern 999999
      ProcessValue <- "86_Times_STEP_MAX_TIME_STP_150"
   TextField "Text field_93" at 295,690 size 75x25; Text 'Step 330'
   IOField "I/O field_81" at 385,690 size 75x25; Authorization "Parameter Change"; FormatPattern 999999
      ProcessValue <- "86_Times_STEP_MAX_TIME_STP_330"
   TextField "Text field_94" at 550,690 size 75x25; Text 'Step 510'
   IOField "I/O field_82" at 640,690 size 75x25; Authorization "Parameter Change"; FormatPattern 999999
      ProcessValue <- "86_Times_STEP_MAX_TIME_STP_510"
   TextField "Text field_97" at 40,725 size 75x25; Text 'Step 160'
   IOField "I/O field_85" at 130,725 size 75x25; Authorization "Parameter Change"; FormatPattern 999999
      ProcessValue <- "86_Times_STEP_MAX_TIME_STP_160"
   TextField "Text field_98" at 295,725 size 75x25; Text 'Step 340'
   IOField "I/O field_86" at 385,725 size 75x25; Authorization "Parameter Change"; FormatPattern 999999
      ProcessValue <- "86_Times_STEP_MAX_TIME_STP_340"
   TextField "Text field_99" at 550,725 size 75x25; Text 'Step 520'
   IOField "I/O field_87" at 640,725 size 75x25; Authorization "Parameter Change"; FormatPattern 999999
      ProcessValue <- "86_Times_STEP_MAX_TIME_STP_520"
   Group "Group" at 455,41 size 373x50
   Button "HmiScreenItemData_8" at 469,45 size 355x40; TextOn 'Back'; TextOff 'Text'
   TextField "Screen title" at 455,41 size 373x50; Text 'Screen title'

screen "Inert Gas Conditioning Setup" 1280x800, template "Template"
   on GenerateScreen: "TitleUpdater"()
   Button "HmiScreenItemData_1" at 1,1 size 150x43; TextOn 'Back'; TextOff 'Main Index'
      on Release: ActivateScreen("02 Main Index", 0)
   Button "HmiScreenItemData_3" at 1129,1 size 150x43; TextOn 'I&A Compressor Ok'; TextOff 'Back'
      on Release: function_efd93a16()
   Button "HmiScreenItemData_19" at 675,536 size 570x30; TextOn 'Back'; TextOff 'IGG STEP'; TextList "STEP LIST_GCU"
      ProcessValue <- "100_GCU_AUTO_SEQ_DB_CRNT_STEP"
   AlarmView "Alarm view_1" at 0,777 size 1280x23
   Gauge "Gauge_1" at 210,575 size 200x200; UnitText '%'; CaptionText 'CV 405'
      ProcessValue <- "12_AI_Data_CV_405_SCALED"
   Gauge "Gauge_3" at 5,575 size 200x200; UnitText 'Barg'; CaptionText 'PIT416'
      ProcessValue <- "12_AI_Data_PIT_416_SCALED"
      MaximumValue <- "84_Setpoints_PIT416_HighHigh"
   IOField "I/O field_7" at 575,536 size 90x30; Authorization "Commissioning"; FormatPattern 999; Unit  Step
      ProcessValue <- "100_GCU_AUTO_SEQ_DB_CRNT_STEP"
   Button "HmiScreenItemData_9" at 465,536 size 100x30; TextOn 'Back'; TextOff 'GCU PLC'
   Circle "Circle_2" at 221,271 size 29x29
      Appearance <- "150_GCU_LCL_CNTRL_DB_LCL_CNTRL_ACTV"
   Button "HmiScreenItemData_8" at 44,105 size 230x29; TextOn 'Back'; TextOff 'GCU Mode of Operation'
   Circle "Circle_1" at 221,212 size 29x29
      Appearance <- "82_To_HMI_CRNT_MODE_GCU"
   Button "HmiScreenItemData_4" at 50,202 size 150x51; TextOn 'Back'; TextOff 'Manual'; Authorization "Operating Mode"
      on Press: function_b14e0dd5("80_From_HMI_Request_Manual", 0); ResetBit("150_GCU_LCL_CNTRL_DB_LCL_CNTRL_ACTV")
   Circle "Circle_9" at 221,151 size 29x29
      Appearance <- "82_To_HMI_CRNT_MODE_GCU"
   Button "HmiScreenItemData_23" at 50,141 size 150x51; TextOn 'Back'; TextOff 'Full Auto'; Authorization "Operating Mode"
      on Press: function_b14e0dd5("80_From_HMI_Request_Auto", 0); ResetBit("150_GCU_LCL_CNTRL_DB_LCL_CNTRL_ACTV")
   Button "HmiScreenItemData_7" at 50,263 size 150x51; TextOn 'Back'; TextOff 'Local Auto'; Authorization "User administration"
      on Press: InvertBit("150_GCU_LCL_CNTRL_DB_LCL_CNTRL_ACTV"); function_b14e0dd5("80_From_HMI_Request_Auto", 0); ResetBit("80_From_HMI_Request_Manual")
   TextField "Text field_7" at 325,106 size 282x35; Text 'Recirculating Pump (P-303)'
   Button "Button_7" at 750,110 size 60x25; TextOn 'Alarm'; TextOff 'Service'
      Visibility <- "141_P303_HRS_RUN_DB_SRVC"
      Appearance <- "141_P303_HRS_RUN_DB_SRVC"
   TextField "Text field_14" at 347,179 size 146x20; Text 'Recirculating Pump'
   TextField "Text field_15" at 494,155 size 58x18; Text 'Control'
   TextField "Text field_16" at 569,155 size 64x18; Text 'Running'
   TextField "Text field_1" at 646,154 size 51x18; Text 'Health'
   TextField "Text field_32" at 490,176 size 60x25; Text 'Enabled'
      Appearance <- "14_DQ_DATA_P_303"
   TextField "Text field_2" at 569,176 size 60x25; Text 'Running'
      Appearance <- "10_DI_DATA_P_303_ENBLD"
   Button "Button_2" at 641,176 size 60x25; TextOn 'Alarm'; TextOff 'OK'
      Visibility <- "10_DI_DATA_P_303_OK"
      Appearance <- "10_DI_DATA_P_303_OK"
   GraphicIOField "Graphic I/O field_1" at 750,200 size 60x65; PictureList "Pump Ani"
      ProcessValue <- "10_DI_DATA_P_303_ENBLD"
   Button "HmiScreenItemData_6" at 646,240 size 69x51; TextOn 'Back'; TextOff 'Reset'; Authorization "Operating Mode"
      on Press: function_b14e0dd5("141_P303_HRS_RUN_DB_RST", 0)
   IOField "I/O field_5" at 571,239 size 65x25; FormatPattern 9999; Unit  h
      ProcessValue <- "141_P303_HRS_RUN_DB_SRV_HRS"
   IOField "I/O field_8" at 571,269 size 65x25; Authorization "Commissioning"; FormatPattern 9999; Unit  h
      ProcessValue <- "141_P303_HRS_RUN_DB_SHRS_IP"
   TextField "Text field_11" at 541,241 size 37x20; Text 'Run'
   TextField "Text field_13" at 541,271 size 37x20; Text 'Set'
   TextField "Text field_25" at 584,215 size 100x20; Text 'Service Hour'
   IOField "I/O field_9" at 345,254 size 75x25; FormatPattern 99999; Unit h
      ProcessValue <- "141_P303_HRS_RUN_DB_HRS"
   IOField "I/O field_12" at 422,254 size 40x25; FormatPattern 99; Unit m
      ProcessValue <- "141_P303_HRS_RUN_DB_MINS"
   IOField "I/O field_16" at 464,254 size 40x25; FormatPattern 99; Unit s
      ProcessValue <- "141_P303_HRS_RUN_DB_SECS"
   TextField "Text field_28" at 345,231 size 160x25; Text 'Total Run Time'
   TextField "Text field_3" at 325,325 size 282x35; Text 'Recirculating Pump (P-304)'
   Button "Button_1" at 750,329 size 60x25; TextOn 'Alarm'; TextOff 'Service'
      Appearance <- "142_P304_HRS_RUN_DB_SRVC"
      Visibility <- "142_P304_HRS_RUN_DB_SRVC"
   TextField "Text field_4" at 347,398 size 146x20; Text 'Recirculating Pump'
   TextField "Text field_5" at 494,374 size 58x18; Text 'Control'
   TextField "Text field_6" at 569,374 size 64x18; Text 'Running'
   TextField "Text field_8" at 646,373 size 51x18; Text 'Health'
   TextField "Text field_9" at 490,395 size 60x25; Text 'Enabled'
      Appearance <- "14_DQ_DATA_P_304"
   TextField "Text field_10" at 569,395 size 60x25; Text 'Running'
      Appearance <- "10_DI_DATA_P_304_ENBLD"
   Button "Button_3" at 641,395 size 60x25; TextOn 'Alarm'; TextOff 'OK'
      Appearance <- "10_DI_DATA_P_304_OK"
      Visibility <- "10_DI_DATA_P_304_OK"
   GraphicIOField "Graphic I/O field_2" at 750,419 size 60x65; PictureList "Pump Ani"
      ProcessValue <- "10_DI_DATA_P_304_ENBLD"
   Button "HmiScreenItemData_2" at 646,459 size 69x51; TextOn 'Back'; TextOff 'Reset'; Authorization "Operating Mode"
      on Press: function_b14e0dd5("142_P304_HRS_RUN_DB_RST", 0)
   IOField "I/O field_1" at 571,458 size 65x25; FormatPattern 9999; Unit  h
      ProcessValue <- "142_P304_HRS_RUN_DB_SRV_HRS"
   IOField "I/O field_2" at 571,488 size 65x25; Authorization "Commissioning"; FormatPattern 9999; Unit  h
      ProcessValue <- "142_P304_HRS_RUN_DB_SHRS_IP"
   TextField "Text field_12" at 541,460 size 37x20; Text 'Run'
   TextField "Text field_22" at 541,490 size 37x20; Text 'Set'
   TextField "Text field_23" at 584,434 size 100x20; Text 'Service Hour'
   IOField "I/O field_3" at 345,473 size 75x25; FormatPattern 99999; Unit h
      ProcessValue <- "142_P304_HRS_RUN_DB_HRS"
   IOField "I/O field_4" at 422,473 size 40x25; FormatPattern 99; Unit m
      ProcessValue <- "142_P304_HRS_RUN_DB_MINS"
   IOField "I/O field_6" at 464,473 size 40x25; FormatPattern 99; Unit s
      ProcessValue <- "142_P304_HRS_RUN_DB_SECS"
   TextField "Text field_24" at 345,450 size 160x25; Text 'Total Run Time'
   Circle "Circle_3" at 221,151 size 29x29
      Visibility <- "150_GCU_LCL_CNTRL_DB_LCL_CNTRL_ACTV"
   Circle "Circle_4" at 221,271 size 29x29
      Visibility <- "82_To_HMI_CRNT_MODE_GCU"
   Group "Group" at 455,41 size 373x50
   Button "Button_5" at 50,344 size 210x35; TextOff 'PGC Setpoint Protection'
      on Press: function_efd93a16("PGC Setpoint Protection", 400, 200, -1, -1, 1)
   Button "HmiScreenItemData_10" at 469,45 size 355x40; TextOn 'Back'; TextOff 'Text'
   TextField "Screen title" at 455,41 size 373x50; Text 'Screen title'

